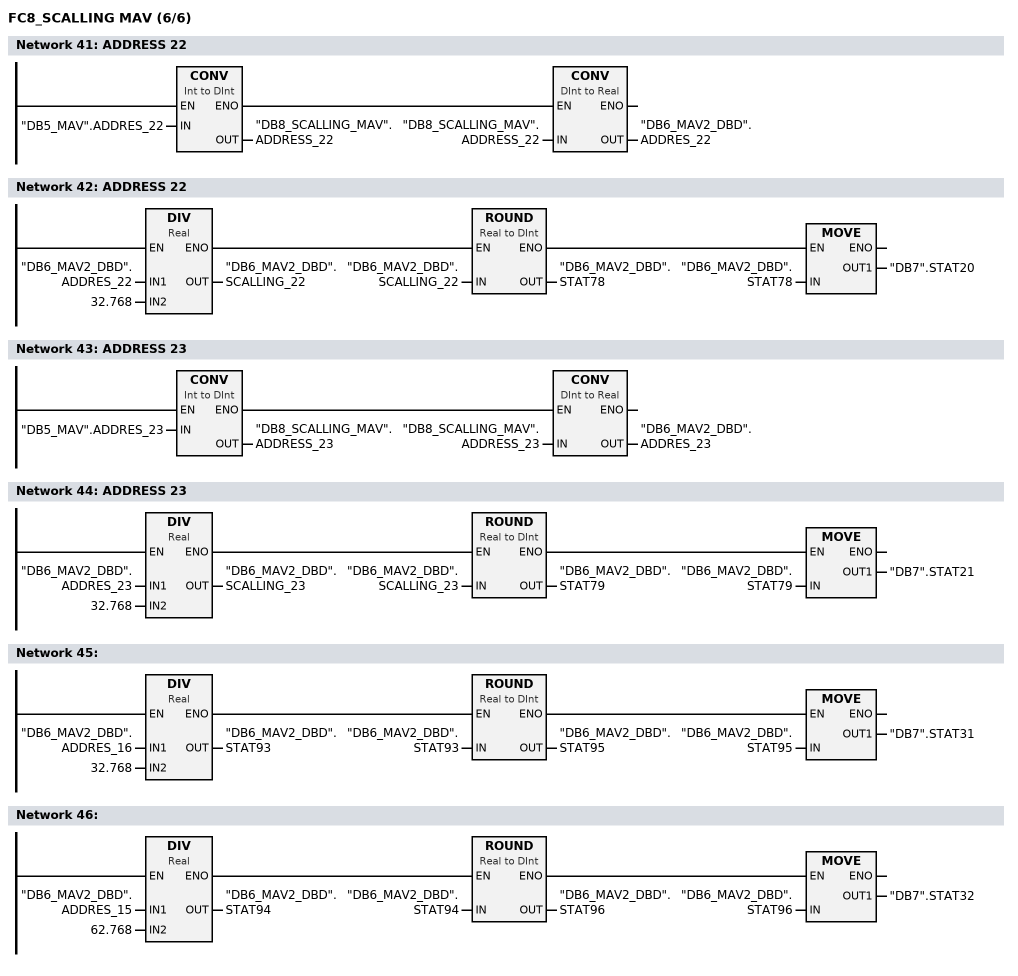
   RUNG wire#powerrail
      { S7_Templates := "[SrcType := Int, DestType := DInt]"; S7_GenerateENO := "TRUE" } Convert(in := "DB5_MAV".ADDRES_22, out => "DB8_SCALLING_MAV".ADDRESS_22)
      { S7_Templates := "[SrcType := DInt, DestType := Real]"; S7_GenerateENO := "TRUE" } Convert(in := "DB8_SCALLING_MAV".ADDRESS_22, out => "DB6_MAV2_DBD".ADDRES_22)
   END_RUNG
   // the same network as SCL:
   // ENO of a box is taken as its EN; it also drops when the box reports an error
   "DB8_SCALLING_MAV".ADDRESS_22 := INT_TO_DINT("DB5_MAV".ADDRES_22);
   "DB6_MAV2_DBD".ADDRES_22 := DINT_TO_REAL("DB8_SCALLING_MAV".ADDRESS_22);
END_REGION

REGION Network 42: ADDRESS 22
   RUNG wire#powerrail
      { S7_Templates := "SrcType := Real"; S7_GenerateENO := "TRUE" } Div(in1 := "DB6_MAV2_DBD".ADDRES_22, in2 := 32.768, out => "DB6_MAV2_DBD".SCALLING_22)
      { S7_Templates := "[SrcType := Real, DestType := DInt]"; S7_GenerateENO := "TRUE" } Round(in := "DB6_MAV2_DBD".SCALLING_22, out => "DB6_MAV2_DBD".STAT78)
      { S7_GenerateENO := "TRUE" } Move(in := "DB6_MAV2_DBD".STAT78, out1 => "DB7".STAT20)
   END_RUNG
   // the same network as SCL:
   // ENO of a box is taken as its EN; it also drops when the box reports an error
   "DB6_MAV2_DBD".SCALLING_22 := "DB6_MAV2_DBD".ADDRES_22 / 32.768;
   "DB6_MAV2_DBD".STAT78 := ROUND("DB6_MAV2_DBD".SCALLING_22);
   "DB7".STAT20 := "DB6_MAV2_DBD".STAT78;
END_REGION

REGION Network 43: ADDRESS 23
   RUNG wire#powerrail
      { S7_Templates := "[SrcType := Int, DestType := DInt]"; S7_GenerateENO := "TRUE" } Convert(in := "DB5_MAV".ADDRES_23, out => "DB8_SCALLING_MAV".ADDRESS_23)
      { S7_Templates := "[SrcType := DInt, DestType := Real]"; S7_GenerateENO := "TRUE" } Convert(in := "DB8_SCALLING_MAV".ADDRESS_23, out => "DB6_MAV2_DBD".ADDRES_23)
   END_RUNG
   // the same network as SCL:
   // ENO of a box is taken as its EN; it also drops when the box reports an error
   "DB8_SCALLING_MAV".ADDRESS_23 := INT_TO_DINT("DB5_MAV".ADDRES_23);
   "DB6_MAV2_DBD".ADDRES_23 := DINT_TO_REAL("DB8_SCALLING_MAV".ADDRESS_23);
END_REGION

REGION Network 44: ADDRESS 23
   RUNG wire#powerrail
      { S7_Templates := "SrcType := Real"; S7_GenerateENO := "TRUE" } Div(in1 := "DB6_MAV2_DBD".ADDRES_23, in2 := 32.768, out => "DB6_MAV2_DBD".SCALLING_23)
      { S7_Templates := "[SrcType := Real, DestType := DInt]"; S7_GenerateENO := "TRUE" } Round(in := "DB6_MAV2_DBD".SCALLING_23, out => "DB6_MAV2_DBD".STAT79)
      { S7_GenerateENO := "TRUE" } Move(in := "DB6_MAV2_DBD".STAT79, out1 => "DB7".STAT21)
   END_RUNG
   // the same network as SCL:
   // ENO of a box is taken as its EN; it also drops when the box reports an error
   "DB6_MAV2_DBD".SCALLING_23 := "DB6_MAV2_DBD".ADDRES_23 / 32.768;
   "DB6_MAV2_DBD".STAT79 := ROUND("DB6_MAV2_DBD".SCALLING_23);
   "DB7".STAT21 := "DB6_MAV2_DBD".STAT79;
END_REGION

REGION Network 45
   RUNG wire#powerrail
      { S7_Templates := "SrcType := Real"; S7_GenerateENO := "TRUE" } Div(in1 := "DB6_MAV2_DBD".ADDRES_16, in2 := 32.768, out => "DB6_MAV2_DBD".STAT93)
      { S7_Templates := "[SrcType := Real, DestType := DInt]"; S7_GenerateENO := "TRUE" } Round(in := "DB6_MAV2_DBD".STAT93, out => "DB6_MAV2_DBD".STAT95)
      { S7_GenerateENO := "TRUE" } Move(in := "DB6_MAV2_DBD".STAT95, out1 => "DB7".STAT31)
   END_RUNG
   // the same network as SCL:
   // ENO of a box is taken as its EN; it also drops when the box reports an error
   "DB6_MAV2_DBD".STAT93 := "DB6_MAV2_DBD".ADDRES_16 / 32.768;
   "DB6_MAV2_DBD".STAT95 := ROUND("DB6_MAV2_DBD".STAT93);
   "DB7".STAT31 := "DB6_MAV2_DBD".STAT95;
END_REGION

REGION Network 46
   RUNG wire#powerrail
      { S7_Templates := "SrcType := Real"; S7_GenerateENO := "TRUE" } Div(in1 := "DB6_MAV2_DBD".ADDRES_15, in2 := 62.768, out => "DB6_MAV2_DBD".STAT94)
      { S7_Templates := "[SrcType := Real, DestType := DInt]"; S7_GenerateENO := "TRUE" } Round(in := "DB6_MAV2_DBD".STAT94, out => "DB6_MAV2_DBD".STAT96)
      { S7_GenerateENO := "TRUE" } Move(in := "DB6_MAV2_DBD".STAT96, out1 => "DB7".STAT32)
   END_RUNG
   // the same network as SCL:
   // ENO of a box is taken as its EN; it also drops when the box reports an error
   "DB6_MAV2_DBD".STAT94 := "DB6_MAV2_DBD".ADDRES_15 / 62.768;
   "DB6_MAV2_DBD".STAT96 := ROUND("DB6_MAV2_DBD".STAT94);
   "DB7".STAT32 := "DB6_MAV2_DBD".STAT96;
END_REGION
END_FUNCTION

FUNCTION "FC9" : Void   // FC9, LAD
{ S7_Optimized_Access := 'FALSE' }
VERSION : 0.1
BEGIN
END_FUNCTION

FUNCTION "FC10_INC_DEC_B" : Void   // FC10, LAD
{ S7_Optimized_Access := 'FALSE' }
VERSION : 0.1
   VAR_INPUT
      Sync : Bool;   // Synchron button
      Sync_SPeed : Real;   // Actual speed reference synchron
      INC : Bool;   // Increase Speed
      DEC : Bool;   // Decrease Speed
   END_VAR
   VAR_IN_OUT
      IO4 : Real;
      SyncSpeed : Real;
      Reff : Int;   // Main Reference value
      SingleSpeed : Real;   // Speed Single Synchron
      IO8 : DInt;
      IO9 : DInt;
   END_VAR
   VAR_TEMP   // added for the SCL form of the ladder/FBD networks
      _w1 : Bool;
   END_VAR
BEGIN

REGION Network 1
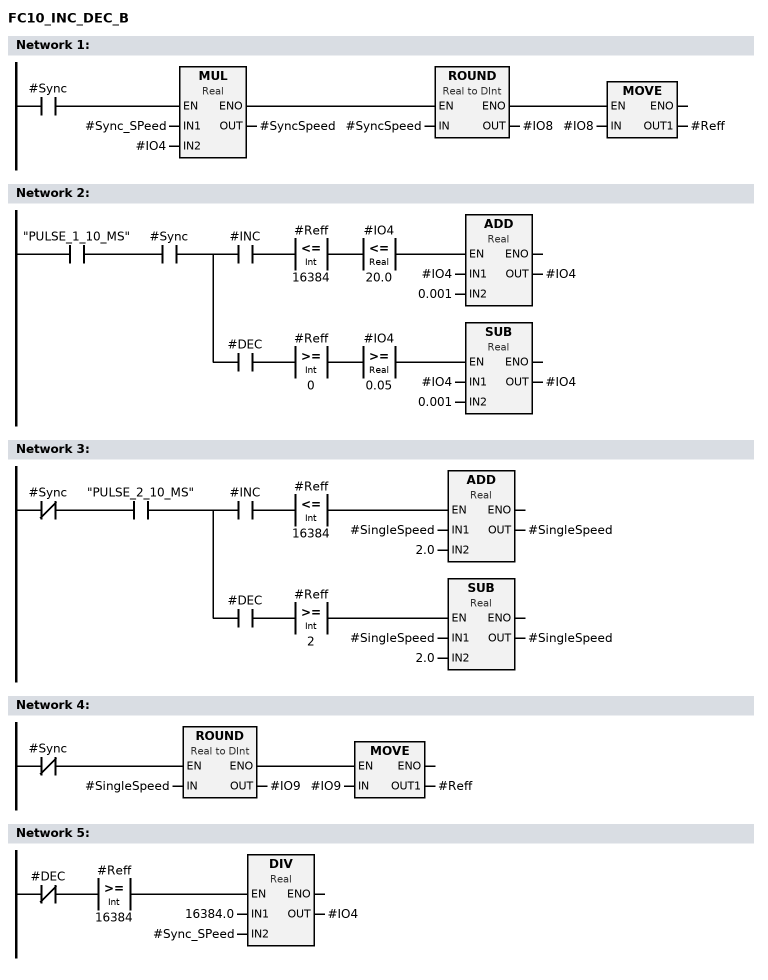
   RUNG wire#powerrail
      Contact( #Sync )
      { S7_Templates := "SrcType := Real"; S7_GenerateENO := "TRUE" } Mul(in1 := #Sync_SPeed, in2 := #IO4, out => #SyncSpeed)
      { S7_Templates := "[SrcType := Real, DestType := DInt]"; S7_GenerateENO := "TRUE" } Round(in := #SyncSpeed, out => #IO8)
      { S7_GenerateENO := "TRUE" } Move(in := #IO8, out1 => #Reff)
   END_RUNG
   // the same network as SCL:
   // ENO of a box is taken as its EN; it also drops when the box reports an error
   IF #Sync THEN
       #SyncSpeed := #Sync_SPeed * #IO4;
       #IO8 := ROUND(#SyncSpeed);
       #Reff := #IO8;
   END_IF;
END_REGION

REGION Network 2
   RUNG wire#powerrail
      Contact( "PULSE_1_10_MS" )
      Contact( #Sync )
      wire#w1
      Contact( #INC )
      { S7_Templates := "SrcType := Int" } LE_Contact(in1 := #Reff, in2 := 16384)
      { S7_Templates := "SrcType := Real" } LE_Contact(in1 := #IO4, in2 := 20.0)
      { S7_Templates := "SrcType := Real"; S7_GenerateENO := "TRUE" } Add(in1 := #IO4, in2 := 0.001, out => #IO4)
   END_RUNG
   RUNG wire#w1
      Contact( #DEC )
      { S7_Templates := "SrcType := Int" } GE_Contact(in1 := #Reff, in2 := 0)
      { S7_Templates := "SrcType := Real" } GE_Contact(in1 := #IO4, in2 := 0.05)
      { S7_Templates := "SrcType := Real"; S7_GenerateENO := "TRUE" } Sub(in1 := #IO4, in2 := 0.001, out => #IO4)
   END_RUNG
   // the same network as SCL:
   #_w1 := "PULSE_1_10_MS" AND #Sync;
   IF #_w1 AND #INC AND (#Reff <= 16384) AND (#IO4 <= 20.0) THEN #IO4 := #IO4 + 0.001; END_IF;
   IF #_w1 AND #DEC AND (#Reff >= 0) AND (#IO4 >= 0.05) THEN #IO4 := #IO4 - 0.001; END_IF;
END_REGION

REGION Network 3
   RUNG wire#powerrail
      I_Contact( #Sync )
      Contact( "PULSE_2_10_MS" )
      wire#w1
      Contact( #INC )
      { S7_Templates := "SrcType := Int" } LE_Contact(in1 := #Reff, in2 := 16384)
      { S7_Templates := "SrcType := Real"; S7_GenerateENO := "TRUE" } Add(in1 := #SingleSpeed, in2 := 2.0, out => #SingleSpeed)
   END_RUNG
   RUNG wire#w1
      Contact( #DEC )
      { S7_Templates := "SrcType := Int" } GE_Contact(in1 := #Reff, in2 := 2)
      { S7_Templates := "SrcType := Real"; S7_GenerateENO := "TRUE" } Sub(in1 := #SingleSpeed, in2 := 2.0, out => #SingleSpeed)
   END_RUNG
   // the same network as SCL:
   #_w1 := NOT #Sync AND "PULSE_2_10_MS";
   IF #_w1 AND #INC AND (#Reff <= 16384) THEN #SingleSpeed := #SingleSpeed + 2.0; END_IF;
   IF #_w1 AND #DEC AND (#Reff >= 2) THEN #SingleSpeed := #SingleSpeed - 2.0; END_IF;
END_REGION

REGION Network 4
   RUNG wire#powerrail
      I_Contact( #Sync )
      { S7_Templates := "[SrcType := Real, DestType := DInt]"; S7_GenerateENO := "TRUE" } Round(in := #SingleSpeed, out => #IO9)
      { S7_GenerateENO := "TRUE" } Move(in := #IO9, out1 => #Reff)
   END_RUNG
   // the same network as SCL:
   // ENO of a box is taken as its EN; it also drops when the box reports an error
   IF NOT #Sync THEN
       #IO9 := ROUND(#SingleSpeed);
       #Reff := #IO9;
   END_IF;
END_REGION

REGION Network 5
   RUNG wire#powerrail
      I_Contact( #DEC )
      { S7_Templates := "SrcType := Int" } GE_Contact(in1 := #Reff, in2 := 16384)
      { S7_Templates := "SrcType := Real"; S7_GenerateENO := "TRUE" } Div(in1 := 16384.0, in2 := #Sync_SPeed, out => #IO4)
   END_RUNG
   // the same network as SCL:
   IF NOT #DEC AND (#Reff >= 16384) THEN #IO4 := 16384.0 / #Sync_SPeed; END_IF;
END_REGION
END_FUNCTION

FUNCTION "FC11_ALARM_NEW" : Void   // FC11, STL
TITLE = ALARM NEW
{ S7_Optimized_Access := 'FALSE' }
AUTHOR : S4P70
VERSION : 0.1
BEGIN

REGION Network 1: statusWord
         L     "statusWord_profiBus_2":P;
         T     "DB15_ALARM".ALARM_ADDRES_2;
         L     "statusWord_profiBus_3":P;
         T     "DB15_ALARM".ALARM_ADDRES_3;
         L     "statusWord_profiBus_4":P;
         T     "DB15_ALARM".ALARM_ADDRES_4;
         L     "statusWord_profiBus_5":P;
         T     "DB15_ALARM".ALARM_ADDRES_5;
         L     "statusWord_profiBus_6":P;
         T     "DB15_ALARM".ALARM_ADDRES_6;
         L     "statusWord_profiBus_7":P;
         T     "DB15_ALARM".ALARM_ADDRES_7;
         L     "statusWord_profiBus_8":P;
         T     "DB15_ALARM".ALARM_ADDRES_8;
         L     "statusWord_profiBus_9":P;
         T     "DB15_ALARM".ALARM_ADDRES_9;
         L     "statusWord_profiBus_10":P;
         T     "DB15_ALARM".ALARM_ADDRES_10;
         L     "statusWord_profiBus_11":P;
         T     "DB15_ALARM".ALARM_ADDRES_11;
         L     "statusWord_profiBus_12":P;
         T     "DB15_ALARM".ALARM_ADDRES_12;
         L     "statusWord_profiBus_13":P;
         T     "DB15_ALARM".ALARM_ADDRES_13;
         L     "statusWord_profiBus_14":P;
         T     "DB15_ALARM".ALARM_ADDRES_14;
         L     "statusWord_profiBus_15":P;
         T     "DB15_ALARM".ALARM_ADDRES_15;
         L     "statusWord_profiBus_16":P;
         T     "DB15_ALARM".ALARM_ADDRES_16;
         L     "statusWord_profiBus_17":P;
         T     "DB15_ALARM".ALARM_ADDRES_17;
         L     "statusWord_profiBus_18":P;
         T     "DB15_ALARM".ALARM_ADDRES_18;
         L     "statusWord_profiBus_19":P;
         T     "DB15_ALARM".ALARM_ADDRES_19;
         L     "statusWord_profiBus_20":P;
         T     "DB15_ALARM".ALARM_ADDRES_20;
         L     "statusWord_profiBus_21":P;
         T     "DB15_ALARM".ALARM_ADDRES_21;
         L     "statusWord_profiBus_22":P;
         T     "DB15_ALARM".ALARM_ADDRES_22;
         L     "statusWord_profiBus_23":P;
         T     "DB15_ALARM".ALARM_ADDRES_23;
END_REGION

REGION Network 2: PROFIBUS STATUS

         A     "DB16_deviceStates".isState[2];
         =     "profibus addres 2 fault";
         A     "DB16_deviceStates".isState[3];
         =     "profibus addres 3 fault";
         A     "DB16_deviceStates".isState[4];
         =     "profibus addres 4 fault";
         A     "DB16_deviceStates".isState[5];
         =     "profibus addres 5 fault";
         A     "DB16_deviceStates".isState[6];
         =     "profibus addres 6 fault";
         A     "DB16_deviceStates".isState[7];
         =     "profibus addres 7 fault";
         A     "DB16_deviceStates".isState[8];
         =     "profibus addres 8 fault";
         A     "DB16_deviceStates".isState[9];
         =     "profibus addres 9 fault";
         A     "DB16_deviceStates".isState[10];
         =     "profibus addres 10 fault";
         A     "DB16_deviceStates".isState[11];
         =     "profibus addres 11 fault";
         A     "DB16_deviceStates".isState[12];
         =     "profibus addres 12 fault";
         A     "DB16_deviceStates".isState[13];
         =     "profibus addres 13 fault";
         A     "DB16_deviceStates".isState[14];
         =     "profibus addres 14 fault";
         A     "DB16_deviceStates".isState[15];
         =     "profibus addres 15 fault";
         A     "DB16_deviceStates".isState[16];
         =     "profibus addres 16 fault";
         A     "DB16_deviceStates".isState[17];
         =     "profibus addres 17 fault";
         A     "DB16_deviceStates".isState[18];
         =     "profibus addres 18 fault";
         A     "DB16_deviceStates".isState[19];
         =     "profibus addres 19 fault";
         A     "DB16_deviceStates".isState[20];
         =     "profibus addres 20 fault";
         A     "DB16_deviceStates".isState[21];
         =     "profibus addres 21 fault";
         A     "DB16_deviceStates".isState[22];
         =     "profibus addres 22 fault";
         A     "DB16_deviceStates".isState[23];
         =     "profibus addres 23 fault";
END_REGION

REGION Network 3
         A     "SB1";
         =     "EMC PRESSED";
END_REGION
END_FUNCTION

ORGANIZATION_BLOCK "OB1_MAIN"   // OB1, LAD, ProgramCycle
TITLE = MAIN PRG
{ S7_Optimized_Access := 'FALSE' }
VERSION : 0.1
   VAR_TEMP
      TEMP0 : Byte;
      TEMP1 : Byte;
      TEMP2 : Byte;
      TEMP3 : Byte;
      TEMP4 : Byte;
      TEMP5 : Byte;
      TEMP6 : Int;
      TEMP7 : Int;
      TEMP8 : Int;
      TEMP9 : Date_And_Time;
      TEMP10 : Struct
         TEMP11 : Word;
         TEMP12 : Word;
      END_STRUCT;
   END_VAR
   VAR_TEMP   // added for the SCL form of the ladder/FBD networks
      _s5time1 : S5Time;
      _w1 : Bool;
   END_VAR
BEGIN

REGION Network 1: CLOCK M100.0
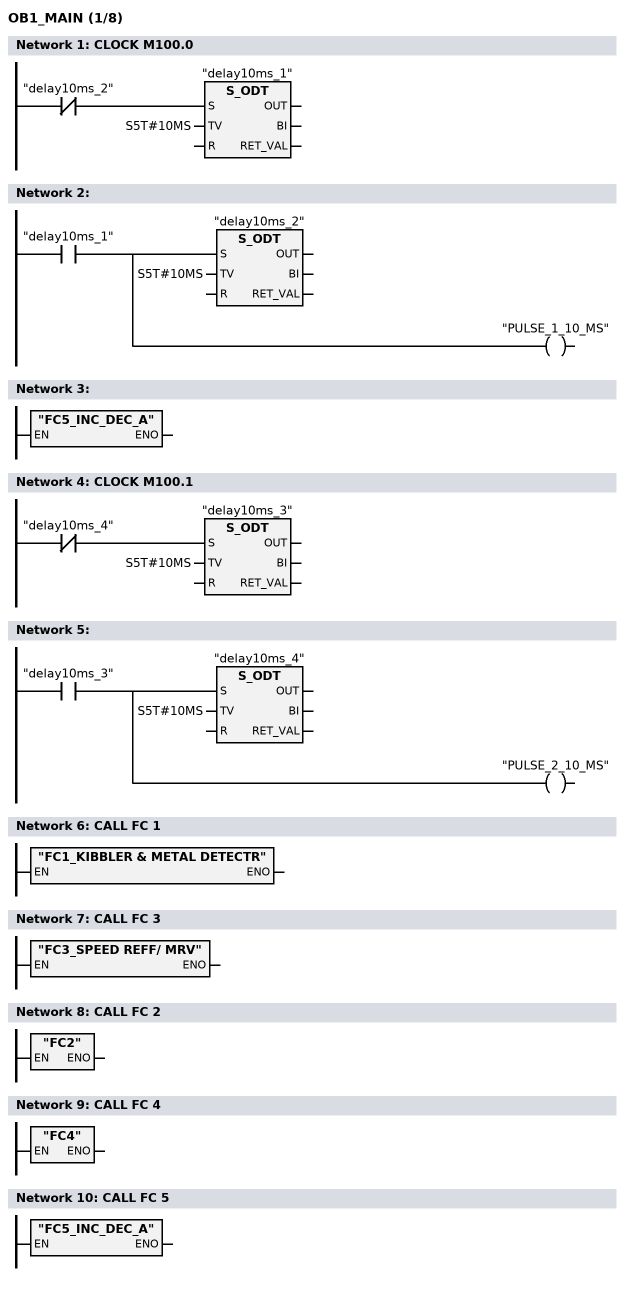
   RUNG wire#powerrail
      I_Contact( "delay10ms_2" )
      S_ODT(T_NO := "delay10ms_1", TV := S5T#10MS, R :=, BI =>, RET_VAL =>)
   END_RUNG
   // the same network as SCL:
   #_s5time1 := S_ODT(T_NO := "delay10ms_1", S := NOT "delay10ms_2", TV := S5T#10MS);
END_REGION

REGION Network 2
   RUNG wire#powerrail
      Contact( "delay10ms_1" )
      wire#w1
      S_ODT(T_NO := "delay10ms_2", TV := S5T#10MS, R :=, BI =>, RET_VAL =>)
   END_RUNG
   RUNG wire#w1
      Coil( "PULSE_1_10_MS" )
   END_RUNG
   // the same network as SCL:
   #_w1 := "delay10ms_1";
   #_s5time1 := S_ODT(T_NO := "delay10ms_2", S := "delay10ms_1", TV := S5T#10MS);
   "PULSE_1_10_MS" := #_w1;
END_REGION

REGION Network 3
   RUNG wire#powerrail
      "FC5_INC_DEC_A"()
   END_RUNG
   // the same network as SCL:
   "FC5_INC_DEC_A"();
END_REGION

REGION Network 4: CLOCK M100.1
   RUNG wire#powerrail
      I_Contact( "delay10ms_4" )
      S_ODT(T_NO := "delay10ms_3", TV := S5T#10MS, R :=, BI =>, RET_VAL =>)
   END_RUNG
   // the same network as SCL:
   #_s5time1 := S_ODT(T_NO := "delay10ms_3", S := NOT "delay10ms_4", TV := S5T#10MS);
END_REGION

REGION Network 5
   RUNG wire#powerrail
      Contact( "delay10ms_3" )
      wire#w1
      S_ODT(T_NO := "delay10ms_4", TV := S5T#10MS, R :=, BI =>, RET_VAL =>)
   END_RUNG
   RUNG wire#w1
      Coil( "PULSE_2_10_MS" )
   END_RUNG
   // the same network as SCL:
   #_w1 := "delay10ms_3";
   #_s5time1 := S_ODT(T_NO := "delay10ms_4", S := "delay10ms_3", TV := S5T#10MS);
   "PULSE_2_10_MS" := #_w1;
END_REGION

REGION Network 6: CALL FC 1
   RUNG wire#powerrail
      "FC1_KIBBLER & METAL DETECTR"()
   END_RUNG
   // the same network as SCL:
   "FC1_KIBBLER & METAL DETECTR"();
END_REGION

REGION Network 7: CALL FC 3
   RUNG wire#powerrail
      "FC3_SPEED REFF/ MRV"()
   END_RUNG
   // the same network as SCL:
   "FC3_SPEED REFF/ MRV"();
END_REGION

REGION Network 8: CALL FC 2
   RUNG wire#powerrail
      "FC2"()
   END_RUNG
   // the same network as SCL:
   "FC2"();
END_REGION

REGION Network 9: CALL FC 4
   RUNG wire#powerrail
      "FC4"()
   END_RUNG
   // the same network as SCL:
   "FC4"();
END_REGION

REGION Network 10: CALL FC 5
   RUNG wire#powerrail
      "FC5_INC_DEC_A"()
   END_RUNG
   // the same network as SCL:
   "FC5_INC_DEC_A"();
END_REGION

REGION Network 11: CALL MAV VLT2800 BLK
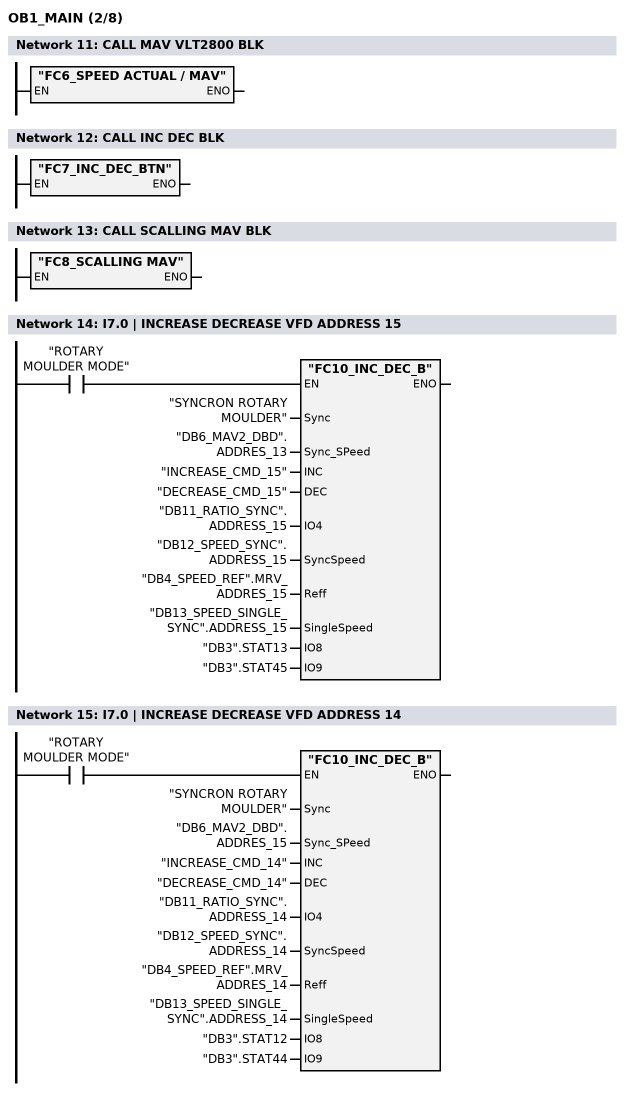
   RUNG wire#powerrail
      "FC6_SPEED ACTUAL / MAV"()
   END_RUNG
   // the same network as SCL:
   "FC6_SPEED ACTUAL / MAV"();
END_REGION

REGION Network 12: CALL INC DEC BLK
   RUNG wire#powerrail
      "FC7_INC_DEC_BTN"()
   END_RUNG
   // the same network as SCL:
   "FC7_INC_DEC_BTN"();
END_REGION

REGION Network 13: CALL SCALLING MAV BLK
   RUNG wire#powerrail
      "FC8_SCALLING MAV"()
   END_RUNG
   // the same network as SCL:
   "FC8_SCALLING MAV"();
END_REGION

REGION Network 14: I7.0 | INCREASE DECREASE VFD ADDRESS 15
   RUNG wire#powerrail
      Contact( "ROTARY MOULDER MODE" )
      "FC10_INC_DEC_B"(Sync := "SYNCRON ROTARY MOULDER", Sync_SPeed := "DB6_MAV2_DBD".ADDRES_13, INC := "INCREASE_CMD_15", DEC := "DECREASE_CMD_15", IO4 := "DB11_RATIO_SYNC".ADDRESS_15, SyncSpeed := "DB12_SPEED_SYNC".ADDRESS_15, Reff := "DB4_SPEED_REF".MRV_ADDRES_15, SingleSpeed := "DB13_SPEED_SINGLE_SYNC".ADDRESS_15, IO8 := "DB3".STAT13, IO9 := "DB3".STAT45)
   END_RUNG
   // the same network as SCL:
   IF "ROTARY MOULDER MODE" THEN
       "FC10_INC_DEC_B"(Sync := "SYNCRON ROTARY MOULDER",
                        Sync_SPeed := "DB6_MAV2_DBD".ADDRES_13,
                        INC := "INCREASE_CMD_15",
                        DEC := "DECREASE_CMD_15",
                        IO4 := "DB11_RATIO_SYNC".ADDRESS_15,
                        SyncSpeed := "DB12_SPEED_SYNC".ADDRESS_15,
                        Reff := "DB4_SPEED_REF".MRV_ADDRES_15,
                        SingleSpeed := "DB13_SPEED_SINGLE_SYNC".ADDRESS_15,
                        IO8 := "DB3".STAT13,
                        IO9 := "DB3".STAT45);
   END_IF;
END_REGION

REGION Network 15: I7.0 | INCREASE DECREASE VFD ADDRESS 14
   RUNG wire#powerrail
      Contact( "ROTARY MOULDER MODE" )
      "FC10_INC_DEC_B"(Sync := "SYNCRON ROTARY MOULDER", Sync_SPeed := "DB6_MAV2_DBD".ADDRES_15, INC := "INCREASE_CMD_14", DEC := "DECREASE_CMD_14", IO4 := "DB11_RATIO_SYNC".ADDRESS_14, SyncSpeed := "DB12_SPEED_SYNC".ADDRESS_14, Reff := "DB4_SPEED_REF".MRV_ADDRES_14, SingleSpeed := "DB13_SPEED_SINGLE_SYNC".ADDRESS_14, IO8 := "DB3".STAT12, IO9 := "DB3".STAT44)
   END_RUNG
   // the same network as SCL:
   IF "ROTARY MOULDER MODE" THEN
       "FC10_INC_DEC_B"(Sync := "SYNCRON ROTARY MOULDER",
                        Sync_SPeed := "DB6_MAV2_DBD".ADDRES_15,
                        INC := "INCREASE_CMD_14",
                        DEC := "DECREASE_CMD_14",
                        IO4 := "DB11_RATIO_SYNC".ADDRESS_14,
                        SyncSpeed := "DB12_SPEED_SYNC".ADDRESS_14,
                        Reff := "DB4_SPEED_REF".MRV_ADDRES_14,
                        SingleSpeed := "DB13_SPEED_SINGLE_SYNC".ADDRESS_14,
                        IO8 := "DB3".STAT12,
                        IO9 := "DB3".STAT44);
   END_IF;
END_REGION

REGION Network 16: I7.0 | INCREASE DECREASE VFD ADDRESS 17
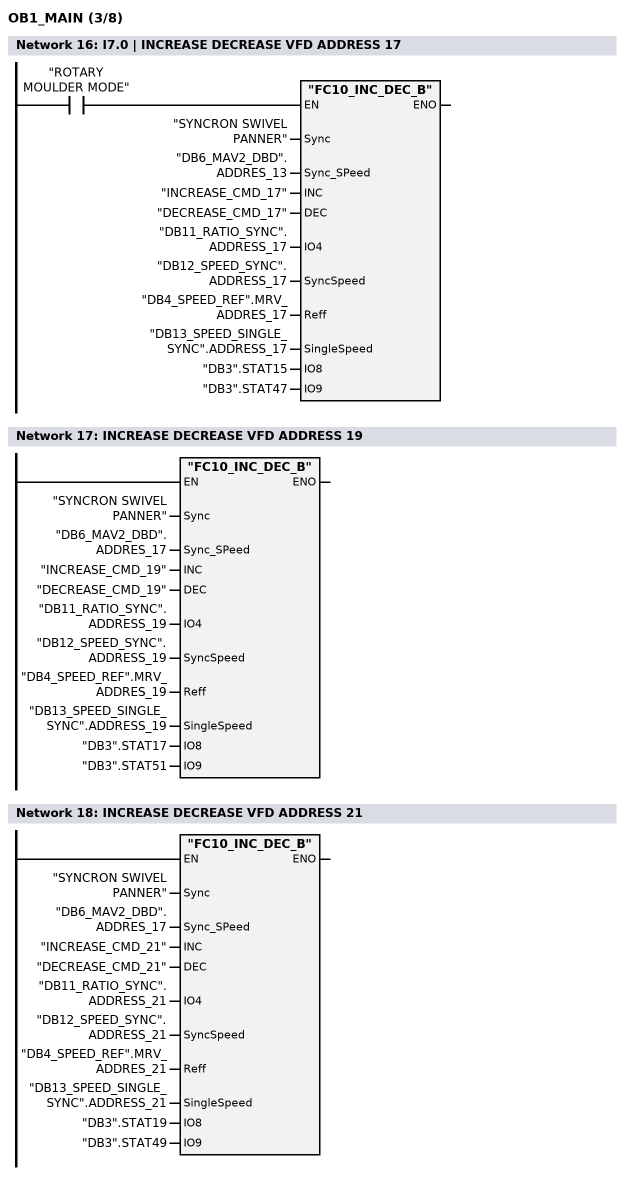
   RUNG wire#powerrail
      Contact( "ROTARY MOULDER MODE" )
      "FC10_INC_DEC_B"(Sync := "SYNCRON SWIVEL PANNER", Sync_SPeed := "DB6_MAV2_DBD".ADDRES_13, INC := "INCREASE_CMD_17", DEC := "DECREASE_CMD_17", IO4 := "DB11_RATIO_SYNC".ADDRESS_17, SyncSpeed := "DB12_SPEED_SYNC".ADDRESS_17, Reff := "DB4_SPEED_REF".MRV_ADDRES_17, SingleSpeed := "DB13_SPEED_SINGLE_SYNC".ADDRESS_17, IO8 := "DB3".STAT15, IO9 := "DB3".STAT47)
   END_RUNG
   // the same network as SCL:
   IF "ROTARY MOULDER MODE" THEN
       "FC10_INC_DEC_B"(Sync := "SYNCRON SWIVEL PANNER",
                        Sync_SPeed := "DB6_MAV2_DBD".ADDRES_13,
                        INC := "INCREASE_CMD_17",
                        DEC := "DECREASE_CMD_17",
                        IO4 := "DB11_RATIO_SYNC".ADDRESS_17,
                        SyncSpeed := "DB12_SPEED_SYNC".ADDRESS_17,
                        Reff := "DB4_SPEED_REF".MRV_ADDRES_17,
                        SingleSpeed := "DB13_SPEED_SINGLE_SYNC".ADDRESS_17,
                        IO8 := "DB3".STAT15,
                        IO9 := "DB3".STAT47);
   END_IF;
END_REGION

REGION Network 17: INCREASE DECREASE VFD ADDRESS 19
   RUNG wire#powerrail
      "FC10_INC_DEC_B"(Sync := "SYNCRON SWIVEL PANNER", Sync_SPeed := "DB6_MAV2_DBD".ADDRES_17, INC := "INCREASE_CMD_19", DEC := "DECREASE_CMD_19", IO4 := "DB11_RATIO_SYNC".ADDRESS_19, SyncSpeed := "DB12_SPEED_SYNC".ADDRESS_19, Reff := "DB4_SPEED_REF".MRV_ADDRES_19, SingleSpeed := "DB13_SPEED_SINGLE_SYNC".ADDRESS_19, IO8 := "DB3".STAT17, IO9 := "DB3".STAT51)
   END_RUNG
   // the same network as SCL:
   "FC10_INC_DEC_B"(Sync := "SYNCRON SWIVEL PANNER",
                    Sync_SPeed := "DB6_MAV2_DBD".ADDRES_17,
                    INC := "INCREASE_CMD_19",
                    DEC := "DECREASE_CMD_19",
                    IO4 := "DB11_RATIO_SYNC".ADDRESS_19,
                    SyncSpeed := "DB12_SPEED_SYNC".ADDRESS_19,
                    Reff := "DB4_SPEED_REF".MRV_ADDRES_19,
                    SingleSpeed := "DB13_SPEED_SINGLE_SYNC".ADDRESS_19,
                    IO8 := "DB3".STAT17,
                    IO9 := "DB3".STAT51);
END_REGION

REGION Network 18: INCREASE DECREASE VFD ADDRESS 21
   RUNG wire#powerrail
      "FC10_INC_DEC_B"(Sync := "SYNCRON SWIVEL PANNER", Sync_SPeed := "DB6_MAV2_DBD".ADDRES_17, INC := "INCREASE_CMD_21", DEC := "DECREASE_CMD_21", IO4 := "DB11_RATIO_SYNC".ADDRESS_21, SyncSpeed := "DB12_SPEED_SYNC".ADDRESS_21, Reff := "DB4_SPEED_REF".MRV_ADDRES_21, SingleSpeed := "DB13_SPEED_SINGLE_SYNC".ADDRESS_21, IO8 := "DB3".STAT19, IO9 := "DB3".STAT49)
   END_RUNG
   // the same network as SCL:
   "FC10_INC_DEC_B"(Sync := "SYNCRON SWIVEL PANNER",
                    Sync_SPeed := "DB6_MAV2_DBD".ADDRES_17,
                    INC := "INCREASE_CMD_21",
                    DEC := "DECREASE_CMD_21",
                    IO4 := "DB11_RATIO_SYNC".ADDRESS_21,
                    SyncSpeed := "DB12_SPEED_SYNC".ADDRESS_21,
                    Reff := "DB4_SPEED_REF".MRV_ADDRES_21,
                    SingleSpeed := "DB13_SPEED_SINGLE_SYNC".ADDRESS_21,
                    IO8 := "DB3".STAT19,
                    IO9 := "DB3".STAT49);
END_REGION

REGION Network 19: INCREASE DECREASE VFD ADDRESS 22
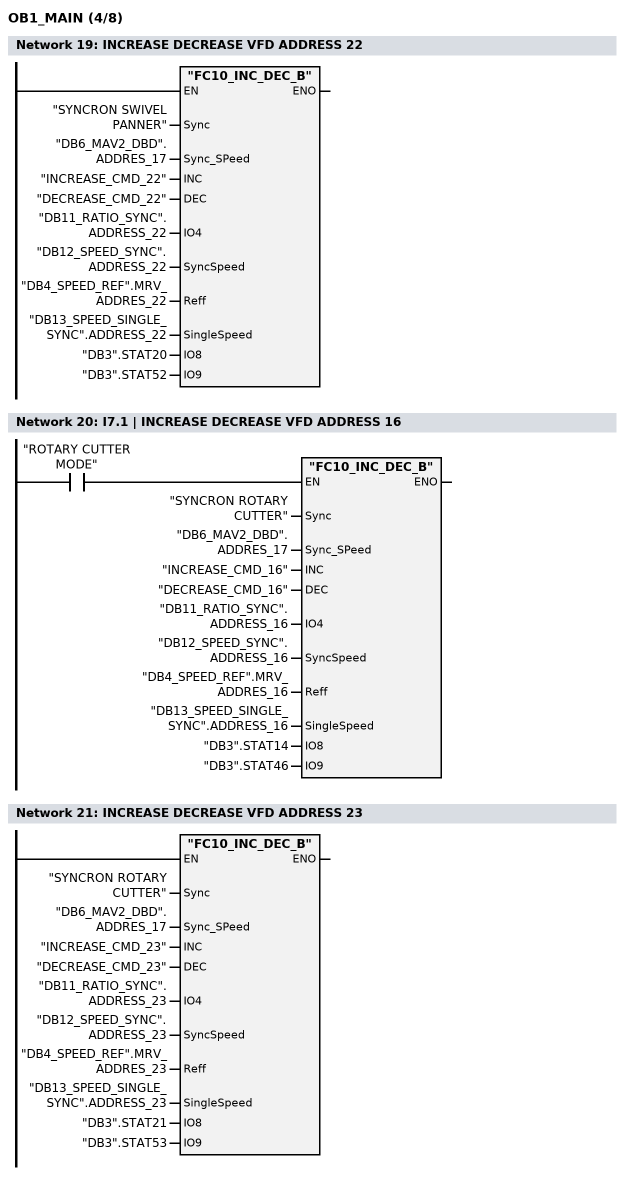
   RUNG wire#powerrail
      "FC10_INC_DEC_B"(Sync := "SYNCRON SWIVEL PANNER", Sync_SPeed := "DB6_MAV2_DBD".ADDRES_17, INC := "INCREASE_CMD_22", DEC := "DECREASE_CMD_22", IO4 := "DB11_RATIO_SYNC".ADDRESS_22, SyncSpeed := "DB12_SPEED_SYNC".ADDRESS_22, Reff := "DB4_SPEED_REF".MRV_ADDRES_22, SingleSpeed := "DB13_SPEED_SINGLE_SYNC".ADDRESS_22, IO8 := "DB3".STAT20, IO9 := "DB3".STAT52)
   END_RUNG
   // the same network as SCL:
   "FC10_INC_DEC_B"(Sync := "SYNCRON SWIVEL PANNER",
                    Sync_SPeed := "DB6_MAV2_DBD".ADDRES_17,
                    INC := "INCREASE_CMD_22",
                    DEC := "DECREASE_CMD_22",
                    IO4 := "DB11_RATIO_SYNC".ADDRESS_22,
                    SyncSpeed := "DB12_SPEED_SYNC".ADDRESS_22,
                    Reff := "DB4_SPEED_REF".MRV_ADDRES_22,
                    SingleSpeed := "DB13_SPEED_SINGLE_SYNC".ADDRESS_22,
                    IO8 := "DB3".STAT20,
                    IO9 := "DB3".STAT52);
END_REGION

REGION Network 20: I7.1 | INCREASE DECREASE VFD ADDRESS 16
   RUNG wire#powerrail
      Contact( "ROTARY CUTTER MODE" )
      "FC10_INC_DEC_B"(Sync := "SYNCRON ROTARY CUTTER", Sync_SPeed := "DB6_MAV2_DBD".ADDRES_17, INC := "INCREASE_CMD_16", DEC := "DECREASE_CMD_16", IO4 := "DB11_RATIO_SYNC".ADDRESS_16, SyncSpeed := "DB12_SPEED_SYNC".ADDRESS_16, Reff := "DB4_SPEED_REF".MRV_ADDRES_16, SingleSpeed := "DB13_SPEED_SINGLE_SYNC".ADDRESS_16, IO8 := "DB3".STAT14, IO9 := "DB3".STAT46)
   END_RUNG
   // the same network as SCL:
   IF "ROTARY CUTTER MODE" THEN
       "FC10_INC_DEC_B"(Sync := "SYNCRON ROTARY CUTTER",
                        Sync_SPeed := "DB6_MAV2_DBD".ADDRES_17,
                        INC := "INCREASE_CMD_16",
                        DEC := "DECREASE_CMD_16",
                        IO4 := "DB11_RATIO_SYNC".ADDRESS_16,
                        SyncSpeed := "DB12_SPEED_SYNC".ADDRESS_16,
                        Reff := "DB4_SPEED_REF".MRV_ADDRES_16,
                        SingleSpeed := "DB13_SPEED_SINGLE_SYNC".ADDRESS_16,
                        IO8 := "DB3".STAT14,
                        IO9 := "DB3".STAT46);
   END_IF;
END_REGION

REGION Network 21: INCREASE DECREASE VFD ADDRESS 23
   RUNG wire#powerrail
      "FC10_INC_DEC_B"(Sync := "SYNCRON ROTARY CUTTER", Sync_SPeed := "DB6_MAV2_DBD".ADDRES_17, INC := "INCREASE_CMD_23", DEC := "DECREASE_CMD_23", IO4 := "DB11_RATIO_SYNC".ADDRESS_23, SyncSpeed := "DB12_SPEED_SYNC".ADDRESS_23, Reff := "DB4_SPEED_REF".MRV_ADDRES_23, SingleSpeed := "DB13_SPEED_SINGLE_SYNC".ADDRESS_23, IO8 := "DB3".STAT21, IO9 := "DB3".STAT53)
   END_RUNG
   // the same network as SCL:
   "FC10_INC_DEC_B"(Sync := "SYNCRON ROTARY CUTTER",
                    Sync_SPeed := "DB6_MAV2_DBD".ADDRES_17,
                    INC := "INCREASE_CMD_23",
                    DEC := "DECREASE_CMD_23",
                    IO4 := "DB11_RATIO_SYNC".ADDRESS_23,
                    SyncSpeed := "DB12_SPEED_SYNC".ADDRESS_23,
                    Reff := "DB4_SPEED_REF".MRV_ADDRES_23,
                    SingleSpeed := "DB13_SPEED_SINGLE_SYNC".ADDRESS_23,
                    IO8 := "DB3".STAT21,
                    IO9 := "DB3".STAT53);
END_REGION

REGION Network 22: I7.1 | INCREASE DECREASE VFD ADDRESS 12
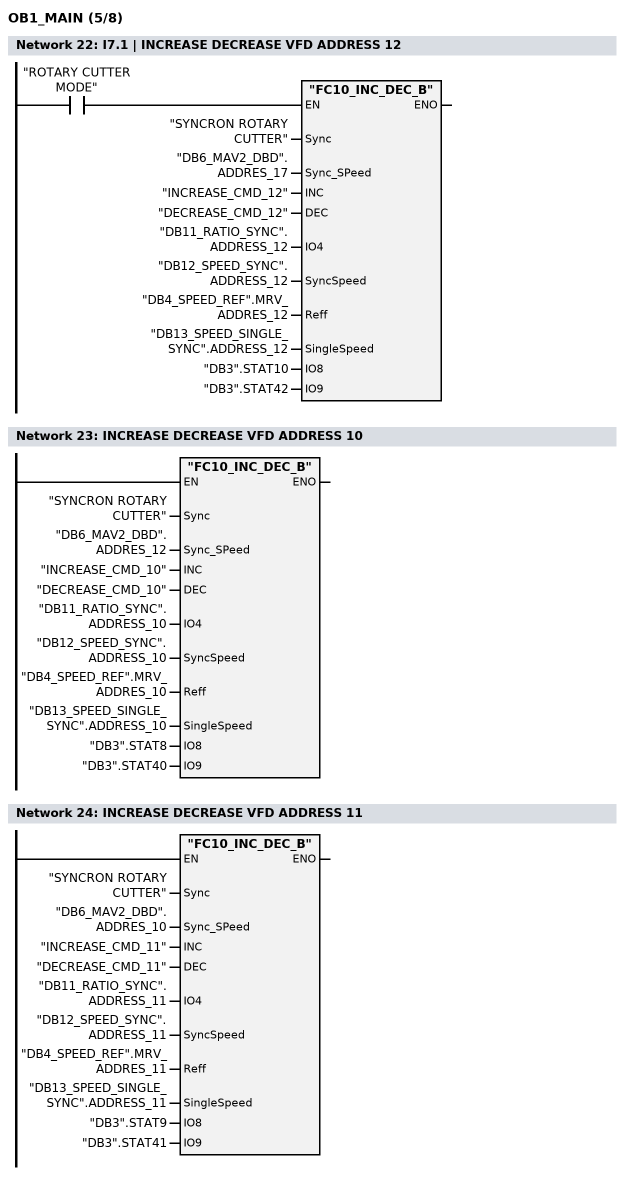
   RUNG wire#powerrail
      Contact( "ROTARY CUTTER MODE" )
      "FC10_INC_DEC_B"(Sync := "SYNCRON ROTARY CUTTER", Sync_SPeed := "DB6_MAV2_DBD".ADDRES_17, INC := "INCREASE_CMD_12", DEC := "DECREASE_CMD_12", IO4 := "DB11_RATIO_SYNC".ADDRESS_12, SyncSpeed := "DB12_SPEED_SYNC".ADDRESS_12, Reff := "DB4_SPEED_REF".MRV_ADDRES_12, SingleSpeed := "DB13_SPEED_SINGLE_SYNC".ADDRESS_12, IO8 := "DB3".STAT10, IO9 := "DB3".STAT42)
   END_RUNG
   // the same network as SCL:
   IF "ROTARY CUTTER MODE" THEN
       "FC10_INC_DEC_B"(Sync := "SYNCRON ROTARY CUTTER",
                        Sync_SPeed := "DB6_MAV2_DBD".ADDRES_17,
                        INC := "INCREASE_CMD_12",
                        DEC := "DECREASE_CMD_12",
                        IO4 := "DB11_RATIO_SYNC".ADDRESS_12,
                        SyncSpeed := "DB12_SPEED_SYNC".ADDRESS_12,
                        Reff := "DB4_SPEED_REF".MRV_ADDRES_12,
                        SingleSpeed := "DB13_SPEED_SINGLE_SYNC".ADDRESS_12,
                        IO8 := "DB3".STAT10,
                        IO9 := "DB3".STAT42);
   END_IF;
END_REGION

REGION Network 23: INCREASE DECREASE VFD ADDRESS 10
   RUNG wire#powerrail
      "FC10_INC_DEC_B"(Sync := "SYNCRON ROTARY CUTTER", Sync_SPeed := "DB6_MAV2_DBD".ADDRES_12, INC := "INCREASE_CMD_10", DEC := "DECREASE_CMD_10", IO4 := "DB11_RATIO_SYNC".ADDRESS_10, SyncSpeed := "DB12_SPEED_SYNC".ADDRESS_10, Reff := "DB4_SPEED_REF".MRV_ADDRES_10, SingleSpeed := "DB13_SPEED_SINGLE_SYNC".ADDRESS_10, IO8 := "DB3".STAT8, IO9 := "DB3".STAT40)
   END_RUNG
   // the same network as SCL:
   "FC10_INC_DEC_B"(Sync := "SYNCRON ROTARY CUTTER",
                    Sync_SPeed := "DB6_MAV2_DBD".ADDRES_12,
                    INC := "INCREASE_CMD_10",
                    DEC := "DECREASE_CMD_10",
                    IO4 := "DB11_RATIO_SYNC".ADDRESS_10,
                    SyncSpeed := "DB12_SPEED_SYNC".ADDRESS_10,
                    Reff := "DB4_SPEED_REF".MRV_ADDRES_10,
                    SingleSpeed := "DB13_SPEED_SINGLE_SYNC".ADDRESS_10,
                    IO8 := "DB3".STAT8,
                    IO9 := "DB3".STAT40);
END_REGION

REGION Network 24: INCREASE DECREASE VFD ADDRESS 11
   RUNG wire#powerrail
      "FC10_INC_DEC_B"(Sync := "SYNCRON ROTARY CUTTER", Sync_SPeed := "DB6_MAV2_DBD".ADDRES_10, INC := "INCREASE_CMD_11", DEC := "DECREASE_CMD_11", IO4 := "DB11_RATIO_SYNC".ADDRESS_11, SyncSpeed := "DB12_SPEED_SYNC".ADDRESS_11, Reff := "DB4_SPEED_REF".MRV_ADDRES_11, SingleSpeed := "DB13_SPEED_SINGLE_SYNC".ADDRESS_11, IO8 := "DB3".STAT9, IO9 := "DB3".STAT41)
   END_RUNG
   // the same network as SCL:
   "FC10_INC_DEC_B"(Sync := "SYNCRON ROTARY CUTTER",
                    Sync_SPeed := "DB6_MAV2_DBD".ADDRES_10,
                    INC := "INCREASE_CMD_11",
                    DEC := "DECREASE_CMD_11",
                    IO4 := "DB11_RATIO_SYNC".ADDRESS_11,
                    SyncSpeed := "DB12_SPEED_SYNC".ADDRESS_11,
                    Reff := "DB4_SPEED_REF".MRV_ADDRES_11,
                    SingleSpeed := "DB13_SPEED_SINGLE_SYNC".ADDRESS_11,
                    IO8 := "DB3".STAT9,
                    IO9 := "DB3".STAT41);
END_REGION

REGION Network 25: INCREASE DECREASE VFD ADDRESS 8